// TIA Portal project "ScatterExample" (V15.1)

(* hardware
DEVICE "S71500/ET200MP station_1"  S7-1500 station
   slot 0: "Rail_0"  Rack  6ES7 590-1***0-0AA0
   slot 1: "PLC_1"  CPU 1511-1 PN  6ES7 511-1AK01-0AB0  V2.6
      slot 3: "CPU display_1"  6ES7591-1AA00-0AA0
*)

// ===== PLC "PLC_1"  CPU 1511-1 PN =====

TYPE "udt1"
   STRUCT
      x0 : Bool;
      x1 : Bool;
      x2 : Bool;
      x3 : Bool;
      x4 : Bool;
      x5 : Bool;
      x6 : Bool;
      x7 : Bool;
      x10 : Bool;
      x11 : Bool;
      x12 : Bool;
      x13 : Bool;
      x14 : Bool;
      x15 : Bool;
      x16 : Bool;
      x17 : Bool;
   END_STRUCT;
END_TYPE

DATA_BLOCK "db1"   // DB1
{ S7_Optimized_Access := 'TRUE' }
VERSION : 0.1
   VAR
      "b" : Byte;
      w : Word;
      dw : DWord;
      arrX16 : Array[0..15] of Bool;
      arrX8 : Array[0..7] of Bool;
      arrX32 : Array[0..31] of Bool;
      stMyVarible : Struct
         x0 : Bool;
         x1 : Bool;
         x2 : Bool;
         x3 : Bool;
         x4 : Bool;
         x5 : Bool;
         x6 : Bool;
         x7 : Bool;
         x10 : Bool;
         x11 : Bool;
         x12 : Bool;
         x13 : Bool;
         x14 : Bool;
         x15 : Bool;
         x16 : Bool;
         x17 : Bool;
      END_STRUCT;
      udtMyVarible : "udt1";
   END_VAR
BEGIN
END_DATA_BLOCK

FUNCTION "fc1" : Void   // FC1, SCL
{ S7_Optimized_Access := 'TRUE' }
VERSION : 0.1
BEGIN


   //Word to Bool Array
   SCATTER(IN:="db1".w,
           OUT=>"db1".arrX16);

   //Dword to Bool Array
   SCATTER(IN:="db1".dw,
           OUT=>"db1".arrX32);

   //Byte to Bool Array
   SCATTER(IN:="db1".b,
           OUT=>"db1".arrX8);

   //Word to Structure 
   SCATTER(IN:="db1".w,
           OUT=>"db1".stMyVarible);

   //Word to Udt
   SCATTER(IN:="db1".w,
           OUT=>"db1".udtMyVarible);
END_FUNCTION

ORGANIZATION_BLOCK "Main"   // OB1, LAD, ProgramCycle
TITLE = "Main Program Sweep (Cycle)"
{ S7_Optimized_Access := 'TRUE' }
VERSION : 0.1
   VAR_INPUT
      Initial_Call : Bool;   // Initial call of this OB
      Remanence : Bool;   // =True, if remanent data are available
   END_VAR
BEGIN

REGION Network 2
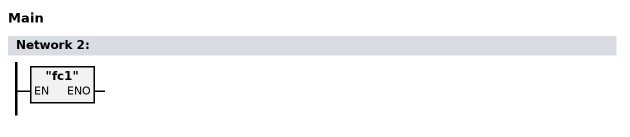
   RUNG wire#powerrail
      "fc1"()
   END_RUNG
   // the same network as SCL:
   "fc1"();
END_REGION
END_ORGANIZATION_BLOCK